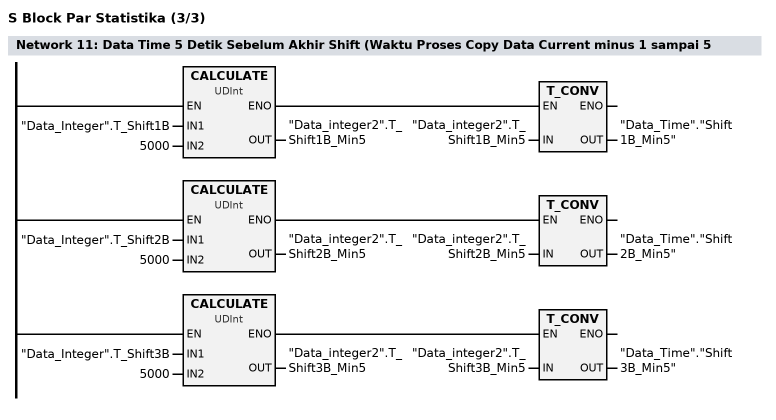
   // ENO of a box is taken as its EN; it also drops when the box reports an error
   "Data_integer2".T_Shift1B_Min5 := "Data_Integer".T_Shift1B-5000;
   "Data_Time"."Shift 1B_Min5" := T_CONV(IN := "Data_integer2".T_Shift1B_Min5);
   "Data_integer2".T_Shift2B_Min5 := "Data_Integer".T_Shift2B-5000;
   "Data_Time"."Shift 2B_Min5" := T_CONV(IN := "Data_integer2".T_Shift2B_Min5);
   "Data_integer2".T_Shift3B_Min5 := "Data_Integer".T_Shift3B-5000;
   "Data_Time"."Shift 3B_Min5" := T_CONV(IN := "Data_integer2".T_Shift3B_Min5);
END_REGION
END_FUNCTION_BLOCK

FUNCTION_BLOCK "S Block Hapus Data"   // FB8, LAD
{ S7_Optimized_Access := 'TRUE' }
VERSION : 0.1
BEGIN

REGION Network 1: Hapus Data Jumlah Sloft Sloft
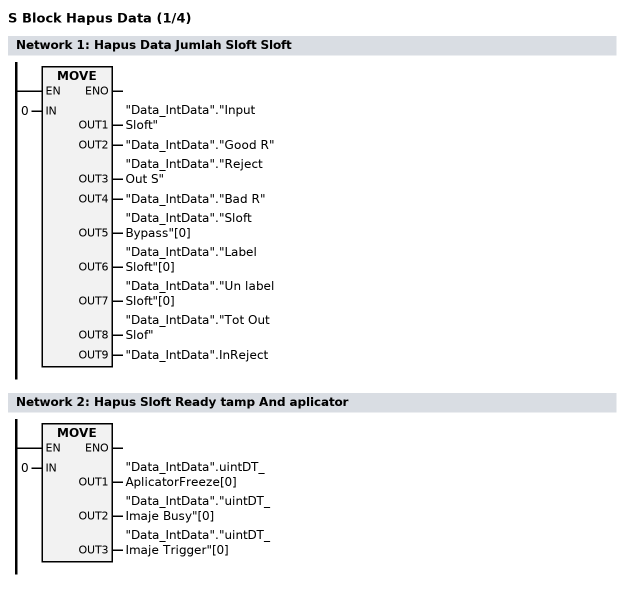
   RUNG wire#powerrail
      { S7_GenerateENO := "TRUE" } Move(in := 0, out1 => "Data_IntData"."Input Sloft", out2 => "Data_IntData"."Good R", out3 => "Data_IntData"."Reject Out S", out4 => "Data_IntData"."Bad R", out5 => "Data_IntData"."Sloft Bypass"[0], out6 => "Data_IntData"."Label Sloft"[0], out7 => "Data_IntData"."Un label Sloft"[0], out8 => "Data_IntData"."Tot Out Slof", out9 => "Data_IntData".InReject)
   END_RUNG
   // the same network as SCL:
   "Data_IntData"."Input Sloft" := 0;
   "Data_IntData"."Good R" := 0;
   "Data_IntData"."Reject Out S" := 0;
   "Data_IntData"."Bad R" := 0;
   "Data_IntData"."Sloft Bypass"[0] := 0;
   "Data_IntData"."Label Sloft"[0] := 0;
   "Data_IntData"."Un label Sloft"[0] := 0;
   "Data_IntData"."Tot Out Slof" := 0;
   "Data_IntData".InReject := 0;
END_REGION

REGION Network 2: Hapus Sloft Ready tamp And aplicator
   RUNG wire#powerrail
      { S7_GenerateENO := "TRUE" } Move(in := 0, out1 => "Data_IntData".uintDT_AplicatorFreeze[0], out2 => "Data_IntData"."uintDT_Imaje Busy"[0], out3 => "Data_IntData"."uintDT_Imaje Trigger"[0])
   END_RUNG
   // the same network as SCL:
   "Data_IntData".uintDT_AplicatorFreeze[0] := 0;
   "Data_IntData"."uintDT_Imaje Busy"[0] := 0;
   "Data_IntData"."uintDT_Imaje Trigger"[0] := 0;
END_REGION

REGION Network 3: Hapus Data Sloft Persen S%
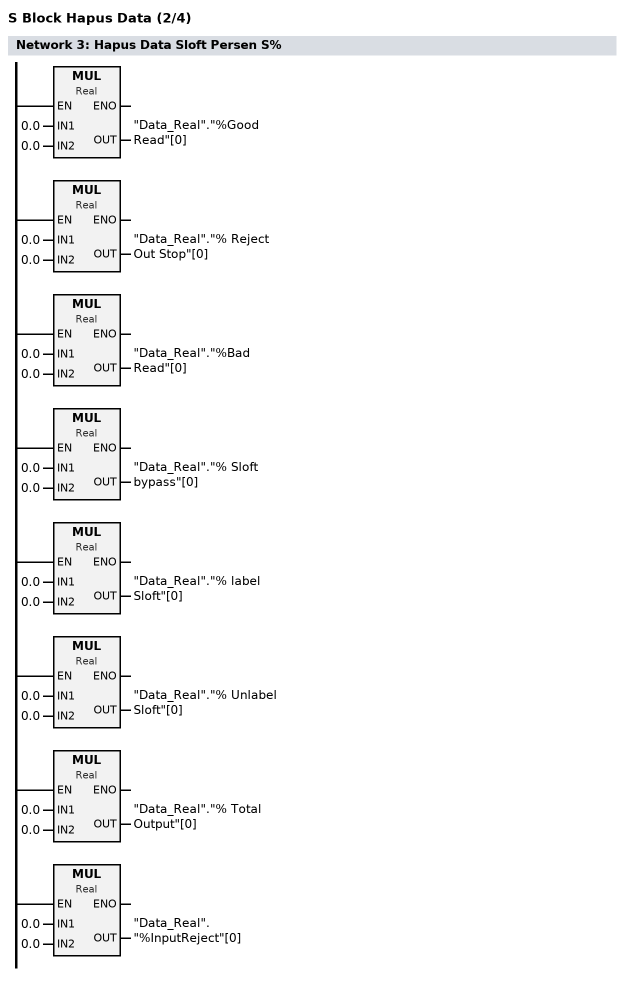
   RUNG wire#powerrail
      { S7_Templates := "SrcType := Real"; S7_GenerateENO := "TRUE" } Mul(in1 := 0.0, in2 := 0.0, out => "Data_Real"."%Good Read"[0])
   END_RUNG
   RUNG wire#powerrail
      { S7_Templates := "SrcType := Real"; S7_GenerateENO := "TRUE" } Mul(in1 := 0.0, in2 := 0.0, out => "Data_Real"."% Reject Out Stop"[0])
   END_RUNG
   RUNG wire#powerrail
      { S7_Templates := "SrcType := Real"; S7_GenerateENO := "TRUE" } Mul(in1 := 0.0, in2 := 0.0, out => "Data_Real"."%Bad Read"[0])
   END_RUNG
   RUNG wire#powerrail
      { S7_Templates := "SrcType := Real"; S7_GenerateENO := "TRUE" } Mul(in1 := 0.0, in2 := 0.0, out => "Data_Real"."% Sloft bypass"[0])
   END_RUNG
   RUNG wire#powerrail
      { S7_Templates := "SrcType := Real"; S7_GenerateENO := "TRUE" } Mul(in1 := 0.0, in2 := 0.0, out => "Data_Real"."% label Sloft"[0])
   END_RUNG
   RUNG wire#powerrail
      { S7_Templates := "SrcType := Real"; S7_GenerateENO := "TRUE" } Mul(in1 := 0.0, in2 := 0.0, out => "Data_Real"."% Unlabel Sloft"[0])
   END_RUNG
   RUNG wire#powerrail
      { S7_Templates := "SrcType := Real"; S7_GenerateENO := "TRUE" } Mul(in1 := 0.0, in2 := 0.0, out => "Data_Real"."% Total Output"[0])
   END_RUNG
   RUNG wire#powerrail
      { S7_Templates := "SrcType := Real"; S7_GenerateENO := "TRUE" } Mul(in1 := 0.0, in2 := 0.0, out => "Data_Real"."%InputReject"[0])
   END_RUNG
   // the same network as SCL:
   "Data_Real"."%Good Read"[0] := 0.0 * 0.0;
   "Data_Real"."% Reject Out Stop"[0] := 0.0 * 0.0;
   "Data_Real"."%Bad Read"[0] := 0.0 * 0.0;
   "Data_Real"."% Sloft bypass"[0] := 0.0 * 0.0;
   "Data_Real"."% label Sloft"[0] := 0.0 * 0.0;
   "Data_Real"."% Unlabel Sloft"[0] := 0.0 * 0.0;
   "Data_Real"."% Total Output"[0] := 0.0 * 0.0;
   "Data_Real"."%InputReject"[0] := 0.0 * 0.0;
END_REGION

REGION Network 4: Hapus Data Time mesin
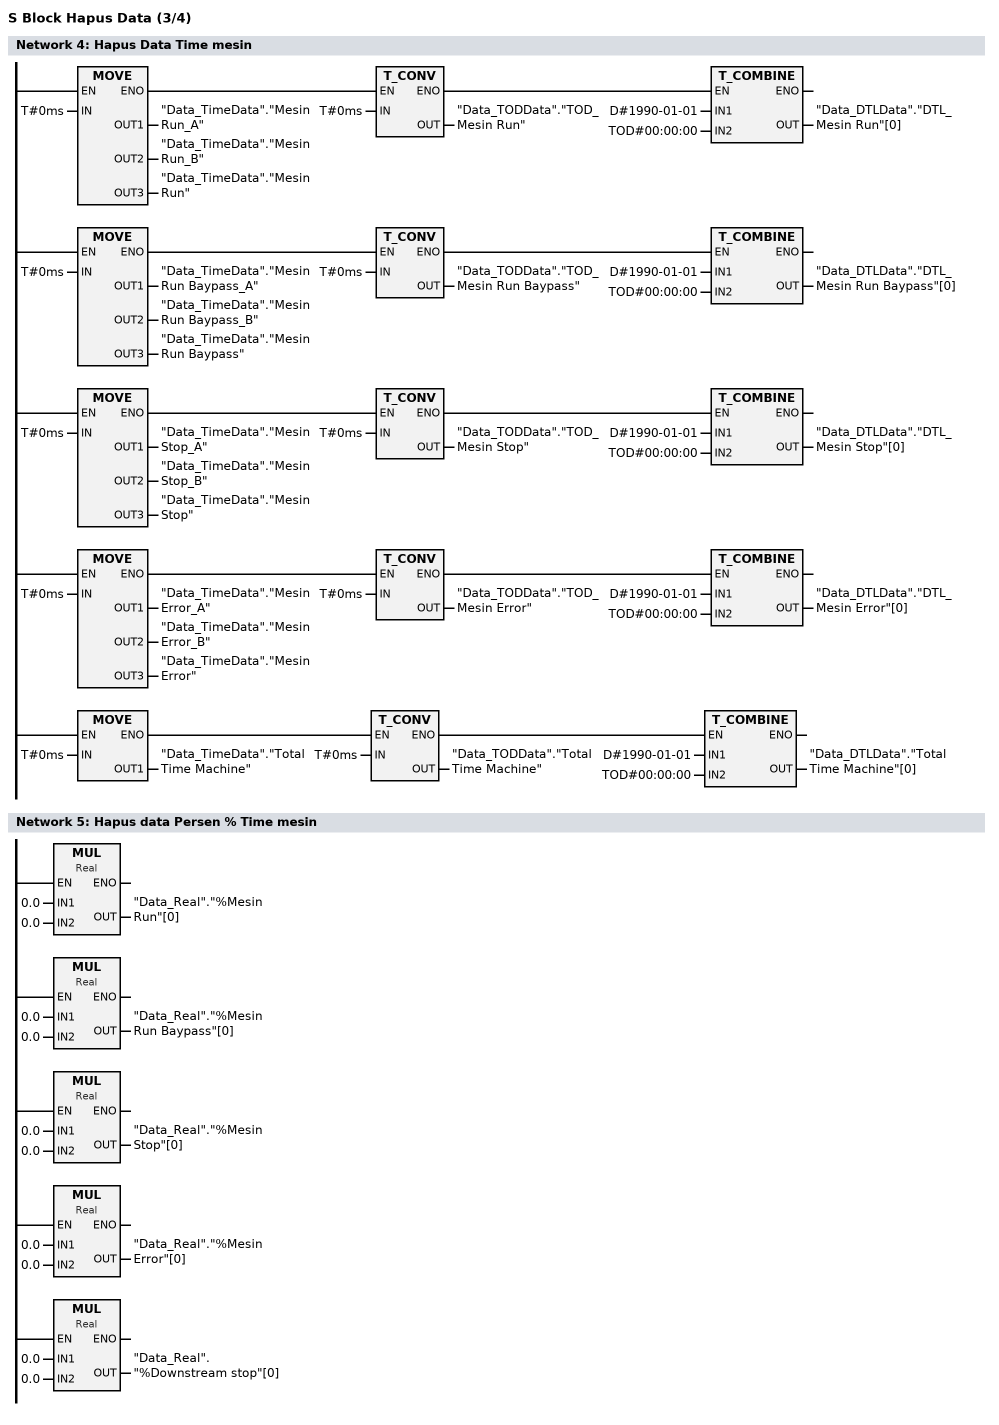
   // ENO of a box is taken as its EN; it also drops when the box reports an error
   "Data_TimeData"."Mesin Run_A" := T#0ms;
   "Data_TimeData"."Mesin Run_B" := T#0ms;
   "Data_TimeData"."Mesin Run" := T#0ms;
   "Data_TODData"."TOD_Mesin Run" := T_CONV(IN := T#0ms);
   "Data_DTLData"."DTL_Mesin Run"[0] := T_COMBINE(IN1 := D#1990-01-01, IN2 := TOD#00:00:00);
   "Data_TimeData"."Mesin Run Baypass_A" := T#0ms;
   "Data_TimeData"."Mesin Run Baypass_B" := T#0ms;
   "Data_TimeData"."Mesin Run Baypass" := T#0ms;
   "Data_TODData"."TOD_Mesin Run Baypass" := T_CONV(IN := T#0ms);
   "Data_DTLData"."DTL_Mesin Run Baypass"[0] := T_COMBINE(IN1 := D#1990-01-01, IN2 := TOD#00:00:00);
   "Data_TimeData"."Mesin Stop_A" := T#0ms;
   "Data_TimeData"."Mesin Stop_B" := T#0ms;
   "Data_TimeData"."Mesin Stop" := T#0ms;
   "Data_TODData"."TOD_Mesin Stop" := T_CONV(IN := T#0ms);
   "Data_DTLData"."DTL_Mesin Stop"[0] := T_COMBINE(IN1 := D#1990-01-01, IN2 := TOD#00:00:00);
   "Data_TimeData"."Mesin Error_A" := T#0ms;
   "Data_TimeData"."Mesin Error_B" := T#0ms;
   "Data_TimeData"."Mesin Error" := T#0ms;
   "Data_TODData"."TOD_Mesin Error" := T_CONV(IN := T#0ms);
   "Data_DTLData"."DTL_Mesin Error"[0] := T_COMBINE(IN1 := D#1990-01-01, IN2 := TOD#00:00:00);
   "Data_TimeData"."Total Time Machine" := T#0ms;
   "Data_TODData"."Total Time Machine" := T_CONV(IN := T#0ms);
   "Data_DTLData"."Total Time Machine"[0] := T_COMBINE(IN1 := D#1990-01-01, IN2 := TOD#00:00:00);
END_REGION

REGION Network 5: Hapus data Persen % Time mesin
   RUNG wire#powerrail
      { S7_Templates := "SrcType := Real"; S7_GenerateENO := "TRUE" } Mul(in1 := 0.0, in2 := 0.0, out => "Data_Real"."%Mesin Run"[0])
   END_RUNG
   RUNG wire#powerrail
      { S7_Templates := "SrcType := Real"; S7_GenerateENO := "TRUE" } Mul(in1 := 0.0, in2 := 0.0, out => "Data_Real"."%Mesin Run Baypass"[0])
   END_RUNG
   RUNG wire#powerrail
      { S7_Templates := "SrcType := Real"; S7_GenerateENO := "TRUE" } Mul(in1 := 0.0, in2 := 0.0, out => "Data_Real"."%Mesin Stop"[0])
   END_RUNG
   RUNG wire#powerrail
      { S7_Templates := "SrcType := Real"; S7_GenerateENO := "TRUE" } Mul(in1 := 0.0, in2 := 0.0, out => "Data_Real"."%Mesin Error"[0])
   END_RUNG
   RUNG wire#powerrail
      { S7_Templates := "SrcType := Real"; S7_GenerateENO := "TRUE" } Mul(in1 := 0.0, in2 := 0.0, out => "Data_Real"."%Downstream stop"[0])
   END_RUNG
   // the same network as SCL:
   "Data_Real"."%Mesin Run"[0] := 0.0 * 0.0;
   "Data_Real"."%Mesin Run Baypass"[0] := 0.0 * 0.0;
   "Data_Real"."%Mesin Stop"[0] := 0.0 * 0.0;
   "Data_Real"."%Mesin Error"[0] := 0.0 * 0.0;
   "Data_Real"."%Downstream stop"[0] := 0.0 * 0.0;
END_REGION

REGION Network 6: Hapus Data Counter Error
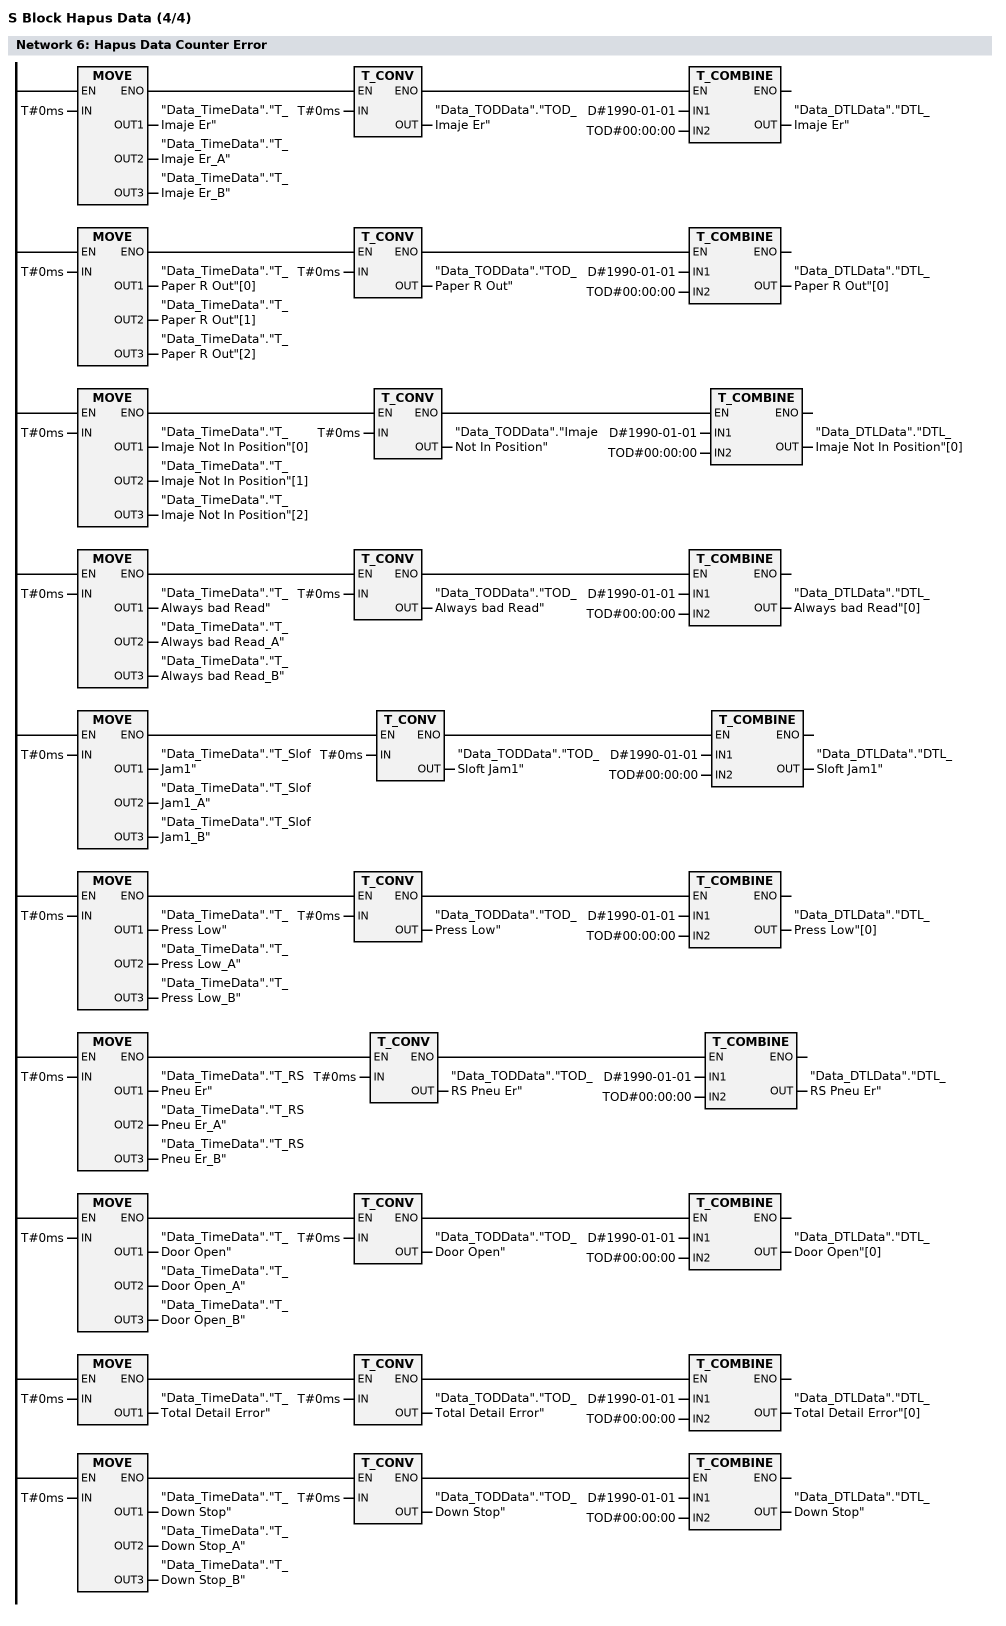
   // ENO of a box is taken as its EN; it also drops when the box reports an error
   "Data_TimeData"."T_Imaje Er" := T#0ms;
   "Data_TimeData"."T_Imaje Er_A" := T#0ms;
   "Data_TimeData"."T_Imaje Er_B" := T#0ms;
   "Data_TODData"."TOD_Imaje Er" := T_CONV(IN := T#0ms);
   "Data_DTLData"."DTL_Imaje Er" := T_COMBINE(IN1 := D#1990-01-01, IN2 := TOD#00:00:00);
   "Data_TimeData"."T_Paper R Out"[0] := T#0ms;
   "Data_TimeData"."T_Paper R Out"[1] := T#0ms;
   "Data_TimeData"."T_Paper R Out"[2] := T#0ms;
   "Data_TODData"."TOD_Paper R Out" := T_CONV(IN := T#0ms);
   "Data_DTLData"."DTL_Paper R Out"[0] := T_COMBINE(IN1 := D#1990-01-01, IN2 := TOD#00:00:00);
   "Data_TimeData"."T_Imaje Not In Position"[0] := T#0ms;
   "Data_TimeData"."T_Imaje Not In Position"[1] := T#0ms;
   "Data_TimeData"."T_Imaje Not In Position"[2] := T#0ms;
   "Data_TODData"."Imaje Not In Position" := T_CONV(IN := T#0ms);
   "Data_DTLData"."DTL_Imaje Not In Position"[0] := T_COMBINE(IN1 := D#1990-01-01, IN2 := TOD#00:00:00);
   "Data_TimeData"."T_Always bad Read" := T#0ms;
   "Data_TimeData"."T_Always bad Read_A" := T#0ms;
   "Data_TimeData"."T_Always bad Read_B" := T#0ms;
   "Data_TODData"."TOD_Always bad Read" := T_CONV(IN := T#0ms);
   "Data_DTLData"."DTL_Always bad Read"[0] := T_COMBINE(IN1 := D#1990-01-01, IN2 := TOD#00:00:00);
   "Data_TimeData"."T_Slof Jam1" := T#0ms;
   "Data_TimeData"."T_Slof Jam1_A" := T#0ms;
   "Data_TimeData"."T_Slof Jam1_B" := T#0ms;
   "Data_TODData"."TOD_Sloft Jam1" := T_CONV(IN := T#0ms);
   "Data_DTLData"."DTL_Sloft Jam1" := T_COMBINE(IN1 := D#1990-01-01, IN2 := TOD#00:00:00);
   "Data_TimeData"."T_Press Low" := T#0ms;
   "Data_TimeData"."T_Press Low_A" := T#0ms;
   "Data_TimeData"."T_Press Low_B" := T#0ms;
   "Data_TODData"."TOD_Press Low" := T_CONV(IN := T#0ms);
   "Data_DTLData"."DTL_Press Low"[0] := T_COMBINE(IN1 := D#1990-01-01, IN2 := TOD#00:00:00);
   "Data_TimeData"."T_RS Pneu Er" := T#0ms;
   "Data_TimeData"."T_RS Pneu Er_A" := T#0ms;
   "Data_TimeData"."T_RS Pneu Er_B" := T#0ms;
   "Data_TODData"."TOD_RS Pneu Er" := T_CONV(IN := T#0ms);
   "Data_DTLData"."DTL_RS Pneu Er" := T_COMBINE(IN1 := D#1990-01-01, IN2 := TOD#00:00:00);
   "Data_TimeData"."T_Door Open" := T#0ms;
   "Data_TimeData"."T_Door Open_A" := T#0ms;
   "Data_TimeData"."T_Door Open_B" := T#0ms;
   "Data_TODData"."TOD_Door Open" := T_CONV(IN := T#0ms);
   "Data_DTLData"."DTL_Door Open"[0] := T_COMBINE(IN1 := D#1990-01-01, IN2 := TOD#00:00:00);
   "Data_TimeData"."T_Total Detail Error" := T#0ms;
   "Data_TODData"."TOD_Total Detail Error" := T_CONV(IN := T#0ms);
   "Data_DTLData"."DTL_Total Detail Error"[0] := T_COMBINE(IN1 := D#1990-01-01, IN2 := TOD#00:00:00);
   "Data_TimeData"."T_Down Stop" := T#0ms;
   "Data_TimeData"."T_Down Stop_A" := T#0ms;
   "Data_TimeData"."T_Down Stop_B" := T#0ms;
   "Data_TODData"."TOD_Down Stop" := T_CONV(IN := T#0ms);
   "Data_DTLData"."DTL_Down Stop" := T_COMBINE(IN1 := D#1990-01-01, IN2 := TOD#00:00:00);
END_REGION
END_FUNCTION_BLOCK

FUNCTION_BLOCK "S Block Current Shift_M1"   // FB9, LAD
TITLE = M1
{ S7_Optimized_Access := 'TRUE' }
VERSION : 0.1
BEGIN

REGION Network 1: Move Date Time M1
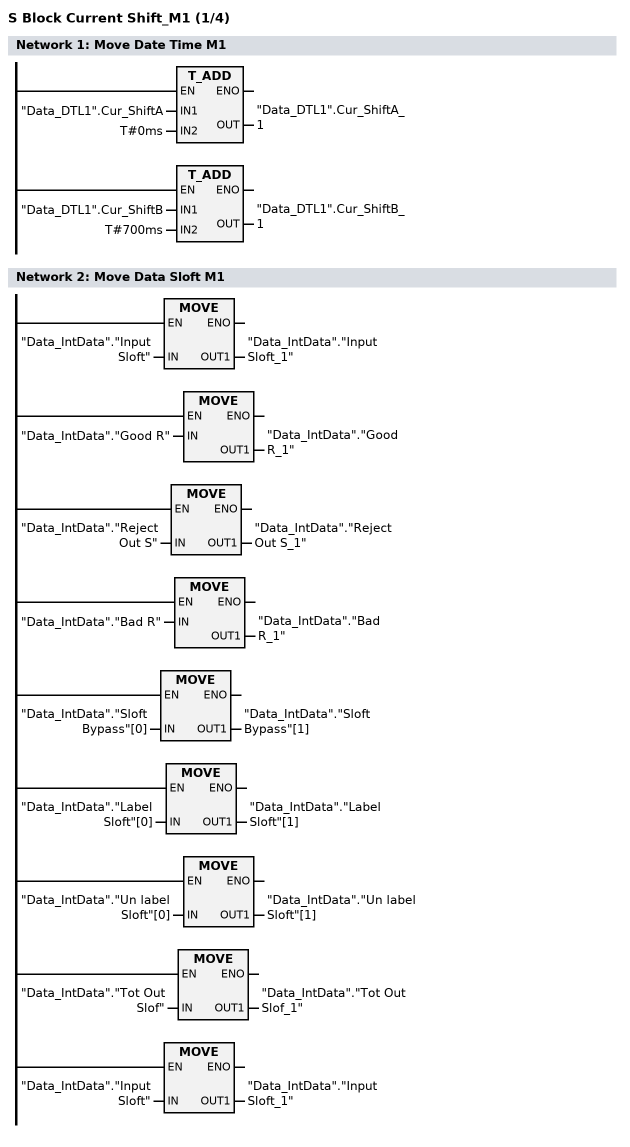
   "Data_DTL1".Cur_ShiftA_1 := T_ADD(IN1 := "Data_DTL1".Cur_ShiftA, IN2 := T#0ms);
   "Data_DTL1".Cur_ShiftB_1 := T_ADD(IN1 := "Data_DTL1".Cur_ShiftB, IN2 := T#700ms);
END_REGION

REGION Network 2: Move Data Sloft M1
   RUNG wire#powerrail
      { S7_GenerateENO := "TRUE" } Move(in := "Data_IntData"."Input Sloft", out1 => "Data_IntData"."Input Sloft_1")
   END_RUNG
   RUNG wire#powerrail
      { S7_GenerateENO := "TRUE" } Move(in := "Data_IntData"."Good R", out1 => "Data_IntData"."Good R_1")
   END_RUNG
   RUNG wire#powerrail
      { S7_GenerateENO := "TRUE" } Move(in := "Data_IntData"."Reject Out S", out1 => "Data_IntData"."Reject Out S_1")
   END_RUNG
   RUNG wire#powerrail
      { S7_GenerateENO := "TRUE" } Move(in := "Data_IntData"."Bad R", out1 => "Data_IntData"."Bad R_1")
   END_RUNG
   RUNG wire#powerrail
      { S7_GenerateENO := "TRUE" } Move(in := "Data_IntData"."Sloft Bypass"[0], out1 => "Data_IntData"."Sloft Bypass"[1])
   END_RUNG
   RUNG wire#powerrail
      { S7_GenerateENO := "TRUE" } Move(in := "Data_IntData"."Label Sloft"[0], out1 => "Data_IntData"."Label Sloft"[1])
   END_RUNG
   RUNG wire#powerrail
      { S7_GenerateENO := "TRUE" } Move(in := "Data_IntData"."Un label Sloft"[0], out1 => "Data_IntData"."Un label Sloft"[1])
   END_RUNG
   RUNG wire#powerrail
      { S7_GenerateENO := "TRUE" } Move(in := "Data_IntData"."Tot Out Slof", out1 => "Data_IntData"."Tot Out Slof_1")
   END_RUNG
   RUNG wire#powerrail
      { S7_GenerateENO := "TRUE" } Move(in := "Data_IntData"."Input Sloft", out1 => "Data_IntData"."Input Sloft_1")
   END_RUNG
   // the same network as SCL:
   "Data_IntData"."Input Sloft_1" := "Data_IntData"."Input Sloft";
   "Data_IntData"."Good R_1" := "Data_IntData"."Good R";
   "Data_IntData"."Reject Out S_1" := "Data_IntData"."Reject Out S";
   "Data_IntData"."Bad R_1" := "Data_IntData"."Bad R";
   "Data_IntData"."Sloft Bypass"[1] := "Data_IntData"."Sloft Bypass"[0];
   "Data_IntData"."Label Sloft"[1] := "Data_IntData"."Label Sloft"[0];
   "Data_IntData"."Un label Sloft"[1] := "Data_IntData"."Un label Sloft"[0];
   "Data_IntData"."Tot Out Slof_1" := "Data_IntData"."Tot Out Slof";
   "Data_IntData"."Input Sloft_1" := "Data_IntData"."Input Sloft";
END_REGION

REGION Network 3: Move Data Sloft Trigger & Aplicator M1
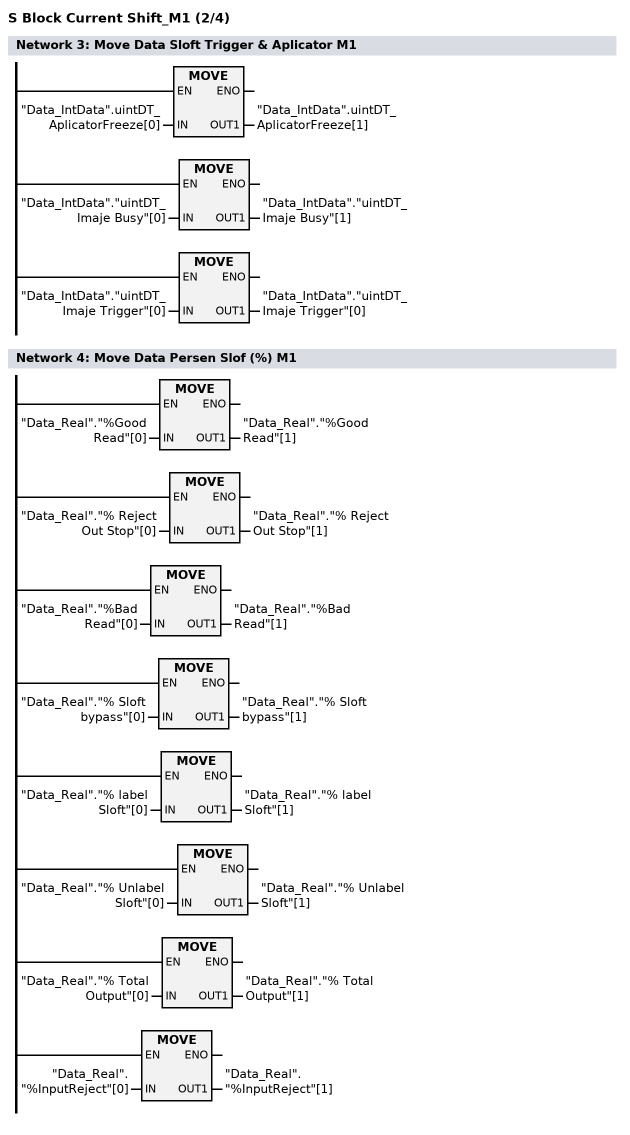
   RUNG wire#powerrail
      { S7_GenerateENO := "TRUE" } Move(in := "Data_IntData".uintDT_AplicatorFreeze[0], out1 => "Data_IntData".uintDT_AplicatorFreeze[1])
   END_RUNG
   RUNG wire#powerrail
      { S7_GenerateENO := "TRUE" } Move(in := "Data_IntData"."uintDT_Imaje Busy"[0], out1 => "Data_IntData"."uintDT_Imaje Busy"[1])
   END_RUNG
   RUNG wire#powerrail
      { S7_GenerateENO := "TRUE" } Move(in := "Data_IntData"."uintDT_Imaje Trigger"[0], out1 => "Data_IntData"."uintDT_Imaje Trigger"[0])
   END_RUNG
   // the same network as SCL:
   "Data_IntData".uintDT_AplicatorFreeze[1] := "Data_IntData".uintDT_AplicatorFreeze[0];
   "Data_IntData"."uintDT_Imaje Busy"[1] := "Data_IntData"."uintDT_Imaje Busy"[0];
   "Data_IntData"."uintDT_Imaje Trigger"[0] := "Data_IntData"."uintDT_Imaje Trigger"[0];
END_REGION

REGION Network 4: Move Data Persen Slof (%) M1
   RUNG wire#powerrail
      { S7_GenerateENO := "TRUE" } Move(in := "Data_Real"."%Good Read"[0], out1 => "Data_Real"."%Good Read"[1])
   END_RUNG
   RUNG wire#powerrail
      { S7_GenerateENO := "TRUE" } Move(in := "Data_Real"."% Reject Out Stop"[0], out1 => "Data_Real"."% Reject Out Stop"[1])
   END_RUNG
   RUNG wire#powerrail
      { S7_GenerateENO := "TRUE" } Move(in := "Data_Real"."%Bad Read"[0], out1 => "Data_Real"."%Bad Read"[1])
   END_RUNG
   RUNG wire#powerrail
      { S7_GenerateENO := "TRUE" } Move(in := "Data_Real"."% Sloft bypass"[0], out1 => "Data_Real"."% Sloft bypass"[1])
   END_RUNG
   RUNG wire#powerrail
      { S7_GenerateENO := "TRUE" } Move(in := "Data_Real"."% label Sloft"[0], out1 => "Data_Real"."% label Sloft"[1])
   END_RUNG
   RUNG wire#powerrail
      { S7_GenerateENO := "TRUE" } Move(in := "Data_Real"."% Unlabel Sloft"[0], out1 => "Data_Real"."% Unlabel Sloft"[1])
   END_RUNG
   RUNG wire#powerrail
      { S7_GenerateENO := "TRUE" } Move(in := "Data_Real"."% Total Output"[0], out1 => "Data_Real"."% Total Output"[1])
   END_RUNG
   RUNG wire#powerrail
      { S7_GenerateENO := "TRUE" } Move(in := "Data_Real"."%InputReject"[0], out1 => "Data_Real"."%InputReject"[1])
   END_RUNG
   // the same network as SCL:
   "Data_Real"."%Good Read"[1] := "Data_Real"."%Good Read"[0];
   "Data_Real"."% Reject Out Stop"[1] := "Data_Real"."% Reject Out Stop"[0];
   "Data_Real"."%Bad Read"[1] := "Data_Real"."%Bad Read"[0];
   "Data_Real"."% Sloft bypass"[1] := "Data_Real"."% Sloft bypass"[0];
   "Data_Real"."% label Sloft"[1] := "Data_Real"."% label Sloft"[0];
   "Data_Real"."% Unlabel Sloft"[1] := "Data_Real"."% Unlabel Sloft"[0];
   "Data_Real"."% Total Output"[1] := "Data_Real"."% Total Output"[0];
   "Data_Real"."%InputReject"[1] := "Data_Real"."%InputReject"[0];
END_REGION

REGION Network 5: Move Data Time Mesin M1
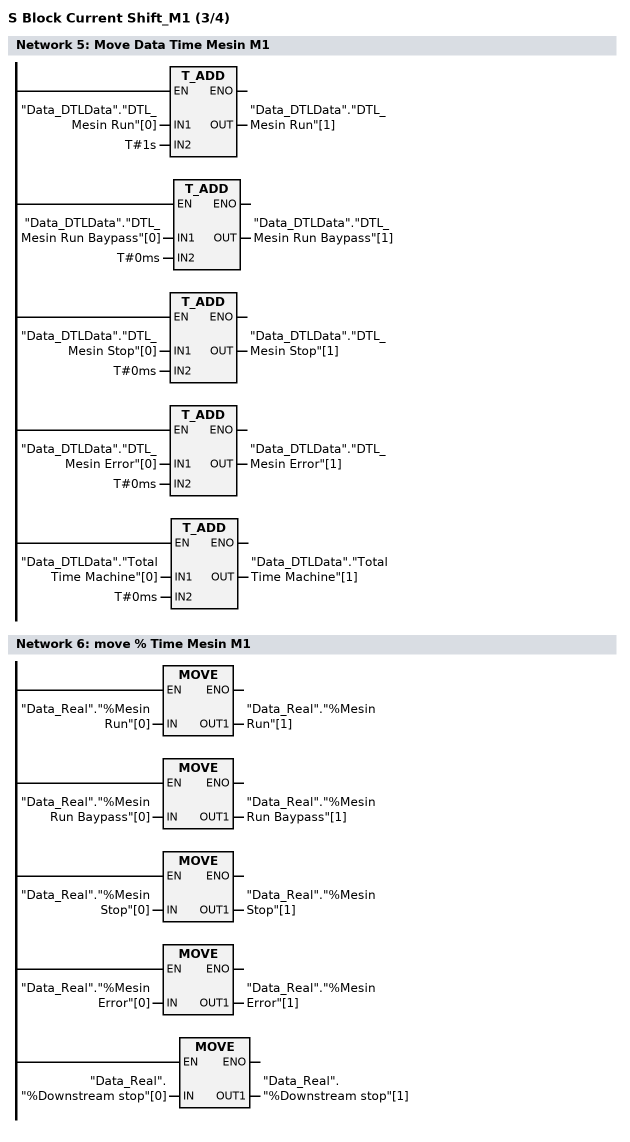
   "Data_DTLData"."DTL_Mesin Run"[1] := T_ADD(IN1 := "Data_DTLData"."DTL_Mesin Run"[0], IN2 := T#1s);
   "Data_DTLData"."DTL_Mesin Run Baypass"[1] := T_ADD(IN1 := "Data_DTLData"."DTL_Mesin Run Baypass"[0],
                           IN2 := T#0ms);
   "Data_DTLData"."DTL_Mesin Stop"[1] := T_ADD(IN1 := "Data_DTLData"."DTL_Mesin Stop"[0], IN2 := T#0ms);
   "Data_DTLData"."DTL_Mesin Error"[1] := T_ADD(IN1 := "Data_DTLData"."DTL_Mesin Error"[0], IN2 := T#0ms);
   "Data_DTLData"."Total Time Machine"[1] := T_ADD(IN1 := "Data_DTLData"."Total Time Machine"[0], IN2 := T#0ms);
END_REGION

REGION Network 6: move % Time Mesin M1
   RUNG wire#powerrail
      { S7_GenerateENO := "TRUE" } Move(in := "Data_Real"."%Mesin Run"[0], out1 => "Data_Real"."%Mesin Run"[1])
   END_RUNG
   RUNG wire#powerrail
      { S7_GenerateENO := "TRUE" } Move(in := "Data_Real"."%Mesin Run Baypass"[0], out1 => "Data_Real"."%Mesin Run Baypass"[1])
   END_RUNG
   RUNG wire#powerrail
      { S7_GenerateENO := "TRUE" } Move(in := "Data_Real"."%Mesin Stop"[0], out1 => "Data_Real"."%Mesin Stop"[1])
   END_RUNG
   RUNG wire#powerrail
      { S7_GenerateENO := "TRUE" } Move(in := "Data_Real"."%Mesin Error"[0], out1 => "Data_Real"."%Mesin Error"[1])
   END_RUNG
   RUNG wire#powerrail
      { S7_GenerateENO := "TRUE" } Move(in := "Data_Real"."%Downstream stop"[0], out1 => "Data_Real"."%Downstream stop"[1])
   END_RUNG
   // the same network as SCL:
   "Data_Real"."%Mesin Run"[1] := "Data_Real"."%Mesin Run"[0];
   "Data_Real"."%Mesin Run Baypass"[1] := "Data_Real"."%Mesin Run Baypass"[0];
   "Data_Real"."%Mesin Stop"[1] := "Data_Real"."%Mesin Stop"[0];
   "Data_Real"."%Mesin Error"[1] := "Data_Real"."%Mesin Error"[0];
   "Data_Real"."%Downstream stop"[1] := "Data_Real"."%Downstream stop"[0];
END_REGION

REGION Network 7: Move Counter Error M1
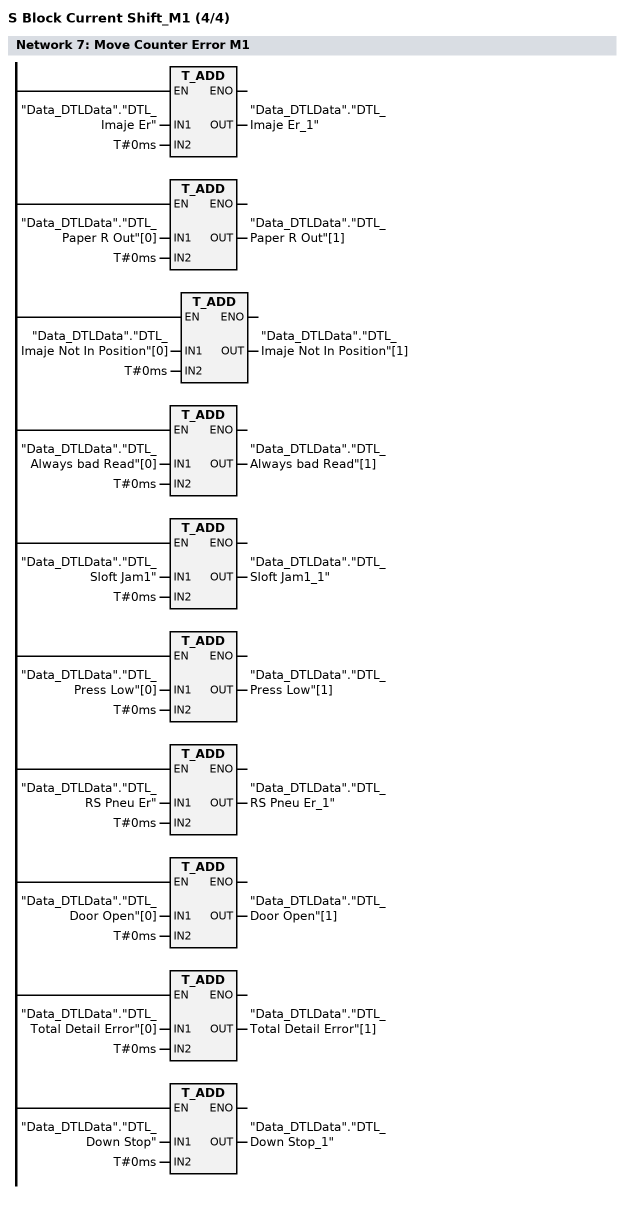
   "Data_DTLData"."DTL_Imaje Er_1" := T_ADD(IN1 := "Data_DTLData"."DTL_Imaje Er", IN2 := T#0ms);
   "Data_DTLData"."DTL_Paper R Out"[1] := T_ADD(IN1 := "Data_DTLData"."DTL_Paper R Out"[0], IN2 := T#0ms);
   "Data_DTLData"."DTL_Imaje Not In Position"[1] := T_ADD(IN1 := "Data_DTLData"."DTL_Imaje Not In Position"[0],
                           IN2 := T#0ms);
   "Data_DTLData"."DTL_Always bad Read"[1] := T_ADD(IN1 := "Data_DTLData"."DTL_Always bad Read"[0],
                           IN2 := T#0ms);
   "Data_DTLData"."DTL_Sloft Jam1_1" := T_ADD(IN1 := "Data_DTLData"."DTL_Sloft Jam1", IN2 := T#0ms);
   "Data_DTLData"."DTL_Press Low"[1] := T_ADD(IN1 := "Data_DTLData"."DTL_Press Low"[0], IN2 := T#0ms);
   "Data_DTLData"."DTL_RS Pneu Er_1" := T_ADD(IN1 := "Data_DTLData"."DTL_RS Pneu Er", IN2 := T#0ms);
   "Data_DTLData"."DTL_Door Open"[1] := T_ADD(IN1 := "Data_DTLData"."DTL_Door Open"[0], IN2 := T#0ms);
   "Data_DTLData"."DTL_Total Detail Error"[1] := T_ADD(IN1 := "Data_DTLData"."DTL_Total Detail Error"[0],
                           IN2 := T#0ms);
   "Data_DTLData"."DTL_Down Stop_1" := T_ADD(IN1 := "Data_DTLData"."DTL_Down Stop", IN2 := T#0ms);
END_REGION
END_FUNCTION_BLOCK

FUNCTION_BLOCK "S Check Range Shift"   // FB10, LAD
{ S7_Optimized_Access := 'TRUE' }
VERSION : 0.1
   VAR_TEMP   // added for the SCL form of the ladder/FBD networks
      _w1 : Bool;
      _w2 : Bool;
      _w3 : Bool;
   END_VAR
BEGIN

REGION Network 1: Check Shift 1
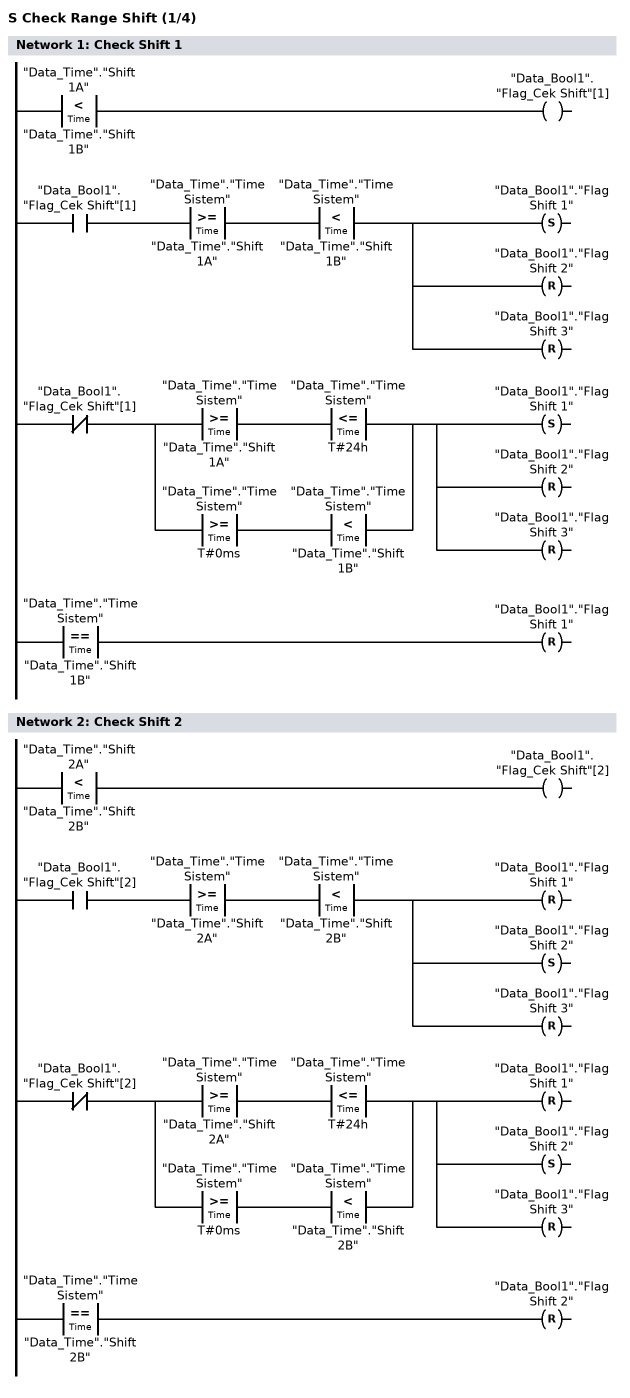
   RUNG wire#powerrail
      { S7_Templates := "SrcType := Time" } LT_Contact(in1 := "Data_Time"."Shift 1A", in2 := "Data_Time"."Shift 1B")
      Coil( "Data_Bool1"."Flag_Cek Shift"[1] )
   END_RUNG
   RUNG wire#powerrail
      Contact( "Data_Bool1"."Flag_Cek Shift"[1] )
      { S7_Templates := "SrcType := Time" } GE_Contact(in1 := "Data_Time"."Time Sistem", in2 := "Data_Time"."Shift 1A")
      { S7_Templates := "SrcType := Time" } LT_Contact(in1 := "Data_Time"."Time Sistem", in2 := "Data_Time"."Shift 1B")
      wire#w1
      S_Coil( "Data_Bool1"."Flag Shift 1" )
   END_RUNG
   RUNG wire#w1
      R_Coil( "Data_Bool1"."Flag Shift 2" )
   END_RUNG
   RUNG wire#w1
      R_Coil( "Data_Bool1"."Flag Shift 3" )
   END_RUNG
   RUNG wire#powerrail
      I_Contact( "Data_Bool1"."Flag_Cek Shift"[1] )
      wire#w2
      { S7_Templates := "SrcType := Time" } GE_Contact(in1 := "Data_Time"."Time Sistem", in2 := "Data_Time"."Shift 1A")
      { S7_Templates := "SrcType := Time" } LE_Contact(in1 := "Data_Time"."Time Sistem", in2 := T#24h)
      wire#w3
      S_Coil( "Data_Bool1"."Flag Shift 1" )
   END_RUNG
   RUNG wire#w2
      { S7_Templates := "SrcType := Time" } GE_Contact(in1 := "Data_Time"."Time Sistem", in2 := T#0ms)
      { S7_Templates := "SrcType := Time" } LT_Contact(in1 := "Data_Time"."Time Sistem", in2 := "Data_Time"."Shift 1B")
   END_RUNG wire#w3
   RUNG wire#w3
      R_Coil( "Data_Bool1"."Flag Shift 2" )
   END_RUNG
   RUNG wire#w3
      R_Coil( "Data_Bool1"."Flag Shift 3" )
   END_RUNG
   RUNG wire#powerrail
      { S7_Templates := "SrcType := Time" } EQ_Contact(in1 := "Data_Time"."Time Sistem", in2 := "Data_Time"."Shift 1B")
      R_Coil( "Data_Bool1"."Flag Shift 1" )
   END_RUNG
   // the same network as SCL:
   "Data_Bool1"."Flag_Cek Shift"[1] := "Data_Time"."Shift 1A" < "Data_Time"."Shift 1B";
   IF "Data_Bool1"."Flag_Cek Shift"[1] AND ("Data_Time"."Time Sistem" >= "Data_Time"."Shift 1A") AND ("Data_Time"."Time Sistem" < "Data_Time"."Shift 1B") THEN
       "Data_Bool1"."Flag Shift 1" := TRUE;
       "Data_Bool1"."Flag Shift 2" := FALSE;
       "Data_Bool1"."Flag Shift 3" := FALSE;
   END_IF;
   IF NOT "Data_Bool1"."Flag_Cek Shift"[1] AND ((("Data_Time"."Time Sistem" >= "Data_Time"."Shift 1A") AND ("Data_Time"."Time Sistem" <= T#24h)) OR (("Data_Time"."Time Sistem" >= T#0ms) AND ("Data_Time"."Time Sistem" < "Data_Time"."Shift 1B"))) THEN
       "Data_Bool1"."Flag Shift 1" := TRUE;
       "Data_Bool1"."Flag Shift 2" := FALSE;
       "Data_Bool1"."Flag Shift 3" := FALSE;
   END_IF;
   IF "Data_Time"."Time Sistem" = "Data_Time"."Shift 1B" THEN "Data_Bool1"."Flag Shift 1" := FALSE; END_IF;
END_REGION

REGION Network 2: Check Shift 2
   RUNG wire#powerrail
      { S7_Templates := "SrcType := Time" } LT_Contact(in1 := "Data_Time"."Shift 2A", in2 := "Data_Time"."Shift 2B")
      Coil( "Data_Bool1"."Flag_Cek Shift"[2] )
   END_RUNG
   RUNG wire#powerrail
      Contact( "Data_Bool1"."Flag_Cek Shift"[2] )
      { S7_Templates := "SrcType := Time" } GE_Contact(in1 := "Data_Time"."Time Sistem", in2 := "Data_Time"."Shift 2A")
      { S7_Templates := "SrcType := Time" } LT_Contact(in1 := "Data_Time"."Time Sistem", in2 := "Data_Time"."Shift 2B")
      wire#w1
      R_Coil( "Data_Bool1"."Flag Shift 1" )
   END_RUNG
   RUNG wire#w1
      S_Coil( "Data_Bool1"."Flag Shift 2" )
   END_RUNG
   RUNG wire#w1
      R_Coil( "Data_Bool1"."Flag Shift 3" )
   END_RUNG
   RUNG wire#powerrail
      I_Contact( "Data_Bool1"."Flag_Cek Shift"[2] )
      wire#w2
      { S7_Templates := "SrcType := Time" } GE_Contact(in1 := "Data_Time"."Time Sistem", in2 := "Data_Time"."Shift 2A")
      { S7_Templates := "SrcType := Time" } LE_Contact(in1 := "Data_Time"."Time Sistem", in2 := T#24h)
      wire#w3
      R_Coil( "Data_Bool1"."Flag Shift 1" )
   END_RUNG
   RUNG wire#w2
      { S7_Templates := "SrcType := Time" } GE_Contact(in1 := "Data_Time"."Time Sistem", in2 := T#0ms)
      { S7_Templates := "SrcType := Time" } LT_Contact(in1 := "Data_Time"."Time Sistem", in2 := "Data_Time"."Shift 2B")
   END_RUNG wire#w3
   RUNG wire#w3
      S_Coil( "Data_Bool1"."Flag Shift 2" )
   END_RUNG
   RUNG wire#w3
      R_Coil( "Data_Bool1"."Flag Shift 3" )
   END_RUNG
   RUNG wire#powerrail
      { S7_Templates := "SrcType := Time" } EQ_Contact(in1 := "Data_Time"."Time Sistem", in2 := "Data_Time"."Shift 2B")
      R_Coil( "Data_Bool1"."Flag Shift 2" )
   END_RUNG
   // the same network as SCL:
   "Data_Bool1"."Flag_Cek Shift"[2] := "Data_Time"."Shift 2A" < "Data_Time"."Shift 2B";
   IF "Data_Bool1"."Flag_Cek Shift"[2] AND ("Data_Time"."Time Sistem" >= "Data_Time"."Shift 2A") AND ("Data_Time"."Time Sistem" < "Data_Time"."Shift 2B") THEN
       "Data_Bool1"."Flag Shift 1" := FALSE;
       "Data_Bool1"."Flag Shift 2" := TRUE;
       "Data_Bool1"."Flag Shift 3" := FALSE;
   END_IF;
   IF NOT "Data_Bool1"."Flag_Cek Shift"[2] AND ((("Data_Time"."Time Sistem" >= "Data_Time"."Shift 2A") AND ("Data_Time"."Time Sistem" <= T#24h)) OR (("Data_Time"."Time Sistem" >= T#0ms) AND ("Data_Time"."Time Sistem" < "Data_Time"."Shift 2B"))) THEN
       "Data_Bool1"."Flag Shift 1" := FALSE;
       "Data_Bool1"."Flag Shift 2" := TRUE;
       "Data_Bool1"."Flag Shift 3" := FALSE;
   END_IF;
   IF "Data_Time"."Time Sistem" = "Data_Time"."Shift 2B" THEN "Data_Bool1"."Flag Shift 2" := FALSE; END_IF;
END_REGION

REGION Network 3: Check Shift 3
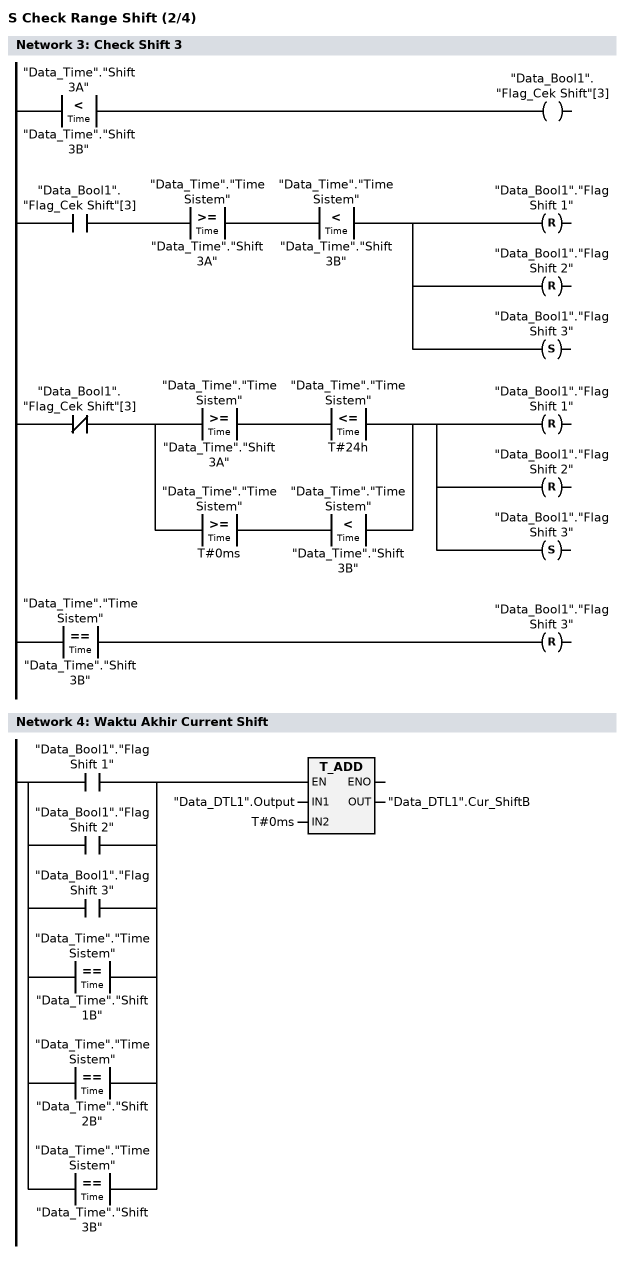
   RUNG wire#powerrail
      { S7_Templates := "SrcType := Time" } LT_Contact(in1 := "Data_Time"."Shift 3A", in2 := "Data_Time"."Shift 3B")
      Coil( "Data_Bool1"."Flag_Cek Shift"[3] )
   END_RUNG
   RUNG wire#powerrail
      Contact( "Data_Bool1"."Flag_Cek Shift"[3] )
      { S7_Templates := "SrcType := Time" } GE_Contact(in1 := "Data_Time"."Time Sistem", in2 := "Data_Time"."Shift 3A")
      { S7_Templates := "SrcType := Time" } LT_Contact(in1 := "Data_Time"."Time Sistem", in2 := "Data_Time"."Shift 3B")
      wire#w1
      R_Coil( "Data_Bool1"."Flag Shift 1" )
   END_RUNG
   RUNG wire#w1
      R_Coil( "Data_Bool1"."Flag Shift 2" )
   END_RUNG
   RUNG wire#w1
      S_Coil( "Data_Bool1"."Flag Shift 3" )
   END_RUNG
   RUNG wire#powerrail
      I_Contact( "Data_Bool1"."Flag_Cek Shift"[3] )
      wire#w2
      { S7_Templates := "SrcType := Time" } GE_Contact(in1 := "Data_Time"."Time Sistem", in2 := "Data_Time"."Shift 3A")
      { S7_Templates := "SrcType := Time" } LE_Contact(in1 := "Data_Time"."Time Sistem", in2 := T#24h)
      wire#w3
      R_Coil( "Data_Bool1"."Flag Shift 1" )
   END_RUNG
   RUNG wire#w2
      { S7_Templates := "SrcType := Time" } GE_Contact(in1 := "Data_Time"."Time Sistem", in2 := T#0ms)
      { S7_Templates := "SrcType := Time" } LT_Contact(in1 := "Data_Time"."Time Sistem", in2 := "Data_Time"."Shift 3B")
   END_RUNG wire#w3
   RUNG wire#w3
      R_Coil( "Data_Bool1"."Flag Shift 2" )
   END_RUNG
   RUNG wire#w3
      S_Coil( "Data_Bool1"."Flag Shift 3" )
   END_RUNG
   RUNG wire#powerrail
      { S7_Templates := "SrcType := Time" } EQ_Contact(in1 := "Data_Time"."Time Sistem", in2 := "Data_Time"."Shift 3B")
      R_Coil( "Data_Bool1"."Flag Shift 3" )
   END_RUNG
   // the same network as SCL:
   "Data_Bool1"."Flag_Cek Shift"[3] := "Data_Time"."Shift 3A" < "Data_Time"."Shift 3B";
   IF "Data_Bool1"."Flag_Cek Shift"[3] AND ("Data_Time"."Time Sistem" >= "Data_Time"."Shift 3A") AND ("Data_Time"."Time Sistem" < "Data_Time"."Shift 3B") THEN
       "Data_Bool1"."Flag Shift 1" := FALSE;
       "Data_Bool1"."Flag Shift 2" := FALSE;
       "Data_Bool1"."Flag Shift 3" := TRUE;
   END_IF;
   IF NOT "Data_Bool1"."Flag_Cek Shift"[3] AND ((("Data_Time"."Time Sistem" >= "Data_Time"."Shift 3A") AND ("Data_Time"."Time Sistem" <= T#24h)) OR (("Data_Time"."Time Sistem" >= T#0ms) AND ("Data_Time"."Time Sistem" < "Data_Time"."Shift 3B"))) THEN
       "Data_Bool1"."Flag Shift 1" := FALSE;
       "Data_Bool1"."Flag Shift 2" := FALSE;
       "Data_Bool1"."Flag Shift 3" := TRUE;
   END_IF;
   IF "Data_Time"."Time Sistem" = "Data_Time"."Shift 3B" THEN "Data_Bool1"."Flag Shift 3" := FALSE; END_IF;
END_REGION

REGION Network 4: Waktu Akhir Current Shift
   IF "Data_Bool1"."Flag Shift 1" OR "Data_Bool1"."Flag Shift 2" OR "Data_Bool1"."Flag Shift 3" OR ("Data_Time"."Time Sistem" = "Data_Time"."Shift 1B") OR ("Data_Time"."Time Sistem" = "Data_Time"."Shift 2B") OR ("Data_Time"."Time Sistem" = "Data_Time"."Shift 3B") THEN
       "Data_DTL1".Cur_ShiftB := T_ADD(IN1 := "Data_DTL1".Output, IN2 := T#0ms);
   END_IF;
END_REGION

REGION Network 5: Waktu Awal Current Shift